(* Logix 5000 project; controller _GigaDiscovery vendor 1 type 14 code 244 rev 35.11; software revision 35.03; part 2 of 23 *)
(* tags used below, declared in another part *)
   Test : DCI_STOP_TEST;

ADD_ON_INSTRUCTION Sfq_Lamp   (* revision 1.0 *)
VAR_INPUT
   Input : BOOL; {required}
END_VAR
VAR_OUTPUT
   LampCoil : BOOL; {access Read Only, visible}
END_VAR
VAR_INPUT
   InputFlt : BOOL; {required}
END_VAR
VAR
   FlsTmr : TIMER := (PRE := 1000); {access None}
END_VAR

ROUTINE Logic   (* ladder *)
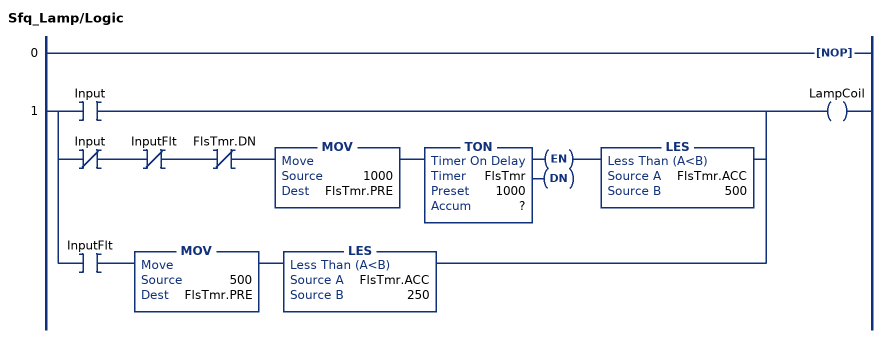
   0: NOP();
   1: [XIC(Input) ,XIO(Input) XIO(InputFlt) XIO(FlsTmr.DN) MOV(1000,FlsTmr.PRE) TON(FlsTmr,?,?) LES(FlsTmr.ACC,500) ,XIC(InputFlt) MOV(500,FlsTmr.PRE) LES(FlsTmr.ACC,250) ]OTE(LampCoil);
END_ROUTINE
END_ADD_ON_INSTRUCTION

ADD_ON_INSTRUCTION Start_AOI   (* revision 1.0 *)
VAR_INPUT
   Start_Ch_1 : BOOL; {required}
   Status_Ch_1 : BOOL; {required}
   Start_Ch_2 : BOOL; {required}
   Status_Ch_2 : BOOL; {required}
   Alarm_Reset : BOOL; {required}
END_VAR
VAR_OUTPUT
   Output : BOOL; {access Read Only, visible}
   Warning : BOOL; {access Read Only, visible}
   Alarm : BOOL; {access Read Only, visible}
   One_Strat_Pb_Pressed : BOOL; {access Read Only}
   Ready : BOOL; {access Read Only}
END_VAR
VAR
   Timer : TIMER[6] := ([0].PRE := 2500, [1].PRE := 2500, [2].PRE := 5000, [3].PRE := 5000, [4].PRE := 5000, [5].PRE := 1000); {access None}
   OS : DINT; {access None}
END_VAR

ROUTINE Logic   (* ladder *)
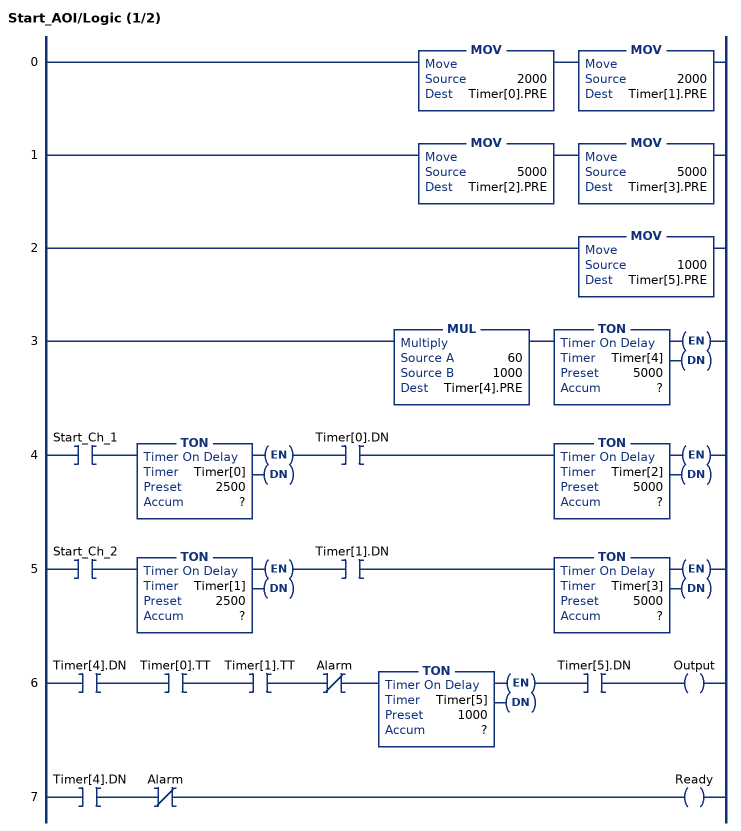
   0: MOV(2000,Timer[0].PRE)MOV(2000,Timer[1].PRE);
   1: MOV(5000,Timer[2].PRE)MOV(5000,Timer[3].PRE);
   2: MOV(1000,Timer[5].PRE);
   3: MUL(60,1000,Timer[4].PRE)TON(Timer[4],?,?);
   4: XIC(Start_Ch_1)TON(Timer[0],?,?)XIC(Timer[0].DN)TON(Timer[2],?,?);
   5: XIC(Start_Ch_2)TON(Timer[1],?,?)XIC(Timer[1].DN)TON(Timer[3],?,?);
   6: XIC(Timer[4].DN)XIC(Timer[0].TT)XIC(Timer[1].TT)XIO(Alarm)TON(Timer[5],?,?)XIC(Timer[5].DN)OTE(Output);
   7: XIC(Timer[4].DN)XIO(Alarm)OTE(Ready);
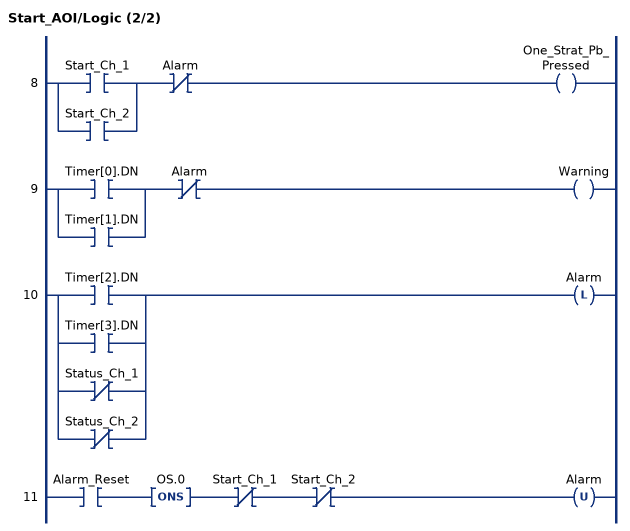
   8: [XIC(Start_Ch_1) ,XIC(Start_Ch_2) ]XIO(Alarm)OTE(One_Strat_Pb_Pressed);
   9: [XIC(Timer[0].DN) ,XIC(Timer[1].DN) ]XIO(Alarm)OTE(Warning);
   10: [XIC(Timer[2].DN) ,XIC(Timer[3].DN) ,XIO(Status_Ch_1) ,XIO(Status_Ch_2) ]OTL(Alarm);
   11: XIC(Alarm_Reset)ONS(OS.0)XIO(Start_Ch_1)XIO(Start_Ch_2)OTU(Alarm);
END_ROUTINE
END_ADD_ON_INSTRUCTION

ADD_ON_INSTRUCTION STD_SCP   (* revision 1.0 *)
VAR_INPUT
   Input : REAL; {required}
   Input_Max : REAL; {required}
   Input_Min : REAL; {required}
END_VAR
VAR_OUTPUT
   Output : REAL; {access Read Only, required}
END_VAR
VAR_INPUT
   Scaled_Max : REAL; {required}
   Scaled_Min : REAL; {required}
END_VAR
VAR
   Rate : REAL;
END_VAR

ROUTINE Logic   (* ladder *)
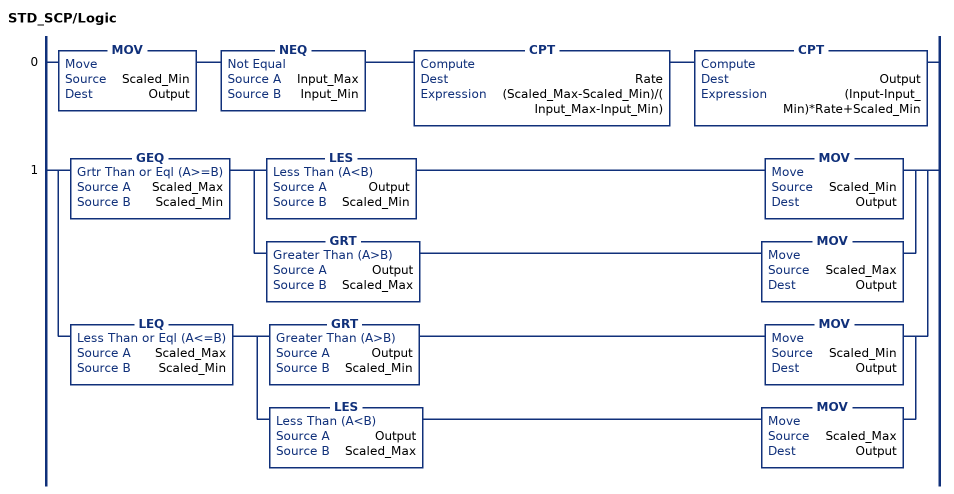
   0: MOV(Scaled_Min,Output)NEQ(Input_Max,Input_Min)CPT(Rate,(Scaled_Max-Scaled_Min)/(Input_Max-Input_Min))CPT(Output,(Input-Input_Min)*Rate+Scaled_Min);
   1: [GEQ(Scaled_Max,Scaled_Min) [LES(Output,Scaled_Min) MOV(Scaled_Min,Output) ,GRT(Output,Scaled_Max) MOV(Scaled_Max,Output) ] ,LEQ(Scaled_Max,Scaled_Min) [GRT(Output,Scaled_Min) MOV(Scaled_Min,Output) ,LES(Output,Scaled_Max) MOV(Scaled_Max,Output) ] ];
END_ROUTINE
END_ADD_ON_INSTRUCTION

ADD_ON_INSTRUCTION Valve_2_pos_monostable   (* revision 1.0 *)
VAR_INPUT
   I_Enable : BOOL; {required}
   FeedBack_Type : BOOL; {required}   // 0 = Equivalent 1 = Reverse
   Discrepancy_Time : DINT; {access None, required}
   I_FeedBack_Data : BOOL; {required}
   I_FeedBack_Status : BOOL; {required}
   I_Output_Status : BOOL; {required}
   I_Fault_Reset : BOOL; {required}
END_VAR
VAR_OUTPUT
   FP : BOOL; {access Read Only, visible}
   O1 : BOOL; {access Read Only, visible}
   O_ERR : DINT; {access Read Only}
END_VAR
VAR
   ON_Delay_Control : TIMER; {access None}
   OFF_Delay_Control : TIMER; {access None}
   Fault_Condiction : BOOL; {access None}
   ONS : BOOL; {access None}
END_VAR

ROUTINE Logic   (* ladder *)
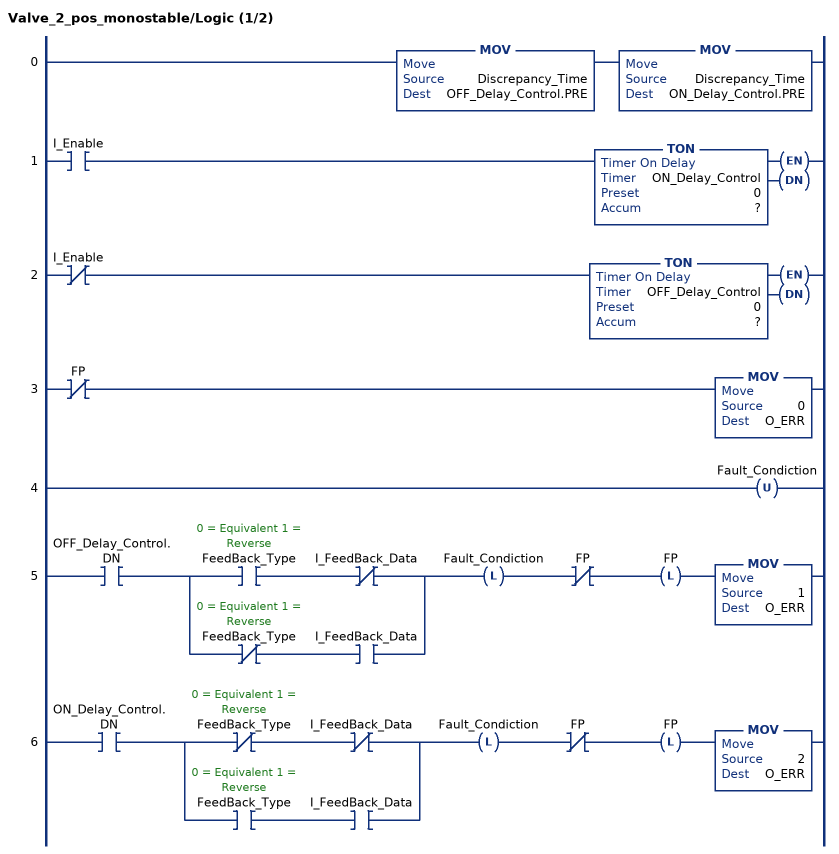
   0: MOV(Discrepancy_Time,OFF_Delay_Control.PRE)MOV(Discrepancy_Time,ON_Delay_Control.PRE);
   1: XIC(I_Enable)TON(ON_Delay_Control,?,?);
   2: XIO(I_Enable)TON(OFF_Delay_Control,?,?);
   3: XIO(FP)MOV(0,O_ERR);
   4: OTU(Fault_Condiction);
   5: XIC(OFF_Delay_Control.DN)[XIC(FeedBack_Type) XIO(I_FeedBack_Data) ,XIO(FeedBack_Type) XIC(I_FeedBack_Data) ]OTL(Fault_Condiction)XIO(FP)OTL(FP)MOV(1,O_ERR);
   6: XIC(ON_Delay_Control.DN)[XIO(FeedBack_Type) XIO(I_FeedBack_Data) ,XIC(FeedBack_Type) XIC(I_FeedBack_Data) ]OTL(Fault_Condiction)XIO(FP)OTL(FP)MOV(2,O_ERR);
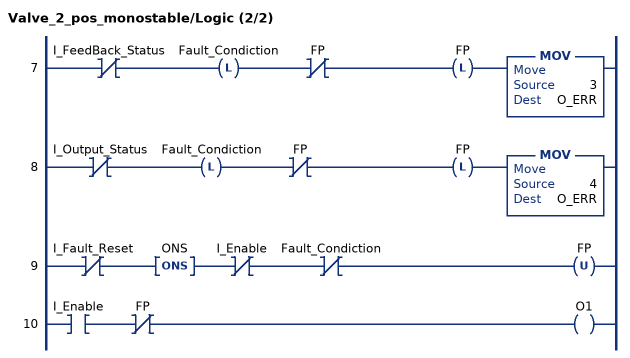
   7: XIO(I_FeedBack_Status)OTL(Fault_Condiction)XIO(FP)OTL(FP)MOV(3,O_ERR);
   8: XIO(I_Output_Status)OTL(Fault_Condiction)XIO(FP)OTL(FP)MOV(4,O_ERR);
   9: XIO(I_Fault_Reset)ONS(ONS)XIO(I_Enable)XIO(Fault_Condiction)OTU(FP);
   10: XIC(I_Enable)XIO(FP)OTE(O1);
END_ROUTINE
END_ADD_ON_INSTRUCTION

VAR_GLOBAL   (* controller tags *)
   Acc_Time : REAL := 0.5;   // T2 Region 2
   All_Rack_Closed_Mem : BOOL := 1;
   All_Rack_Left_Sensor_FP_OFF : BOOL := 1;
   All_Rack_Left_Sensor_O1_OFF : BOOL;
   All_Rack_Right_Sensor_FP_OFF : BOOL := 1;
   All_Rack_Right_Sensor_O1_OFF : BOOL;
   All_Rack_Sensor_OFF : BOOL;
   All_RESTRAINTS_Opened : BOOL;
   Analog_Input_Pos_6 : REAL[8] := ([0] := 0.0061035156, [2] := -0.025939941, [4] := -0.025939941, [6] := -0.0289917);
        [0]   // Lettura tensione Motori 1 - 3 Pilone
        [1]   // Lettura Corrente Motori 1 - 3 Pilone
        [2]   // Lettura tensione Motori 2 - 4 Pilone
        [3]   // Lettura Corrente Motori 2 - 4 Pilone
        [6]   // Lettura tensione Motori 5 - 6 Pilone
        [7]   // Lettura Corrente Motori 5 - 6 Pilone
        [4]   // Lettura tensione Motore Gondola
        [5]   // Lettura Corrente Motore Gondola
   Analog_Output_Pos_5 : REAL[8] := ([4] := 10000.0);
        [4]   // Gondola Torque Limit
        [5]   // Gondola Speed Reference
   Angle_at_Full_Load : REAL := 12.0;
   Angle_at_min_Load : REAL := 14.0;
   Angle_Controll_S_Curve : S_Curve_Calc := (Jerk_Time := 0.5, Accel_Time := 1.0, Jerk_Rate := 300.0, Accel_Rate := 150.0);
   AngleContrl : REAL := 77.39982;
   Auto_Cycle_Step : DINT := 1;
   auto_manual : TIMER := (PRE := 2000);
   Automatic_Cycle_DB : Auto_Cycle[6] := ([1].Pylon_Angle := 120, [1].Cycle_Time_min := 2, [1].Cycle_Time_sec := 25, [1].Gondola_Speed[0] := 20, [1].Gondola_Speed[1] := 70, [1].Gondola_Speed[2] := -75, [1].Gondola_Speed[3] := 50, [1].Gondola_Time[1] := 60, [1].Gondola_Time[2] := 50, [1].Gondola_Time[3] := 20, [2].Pylon_Angle := 90, [2].Cycle_Time_min := 1, [2].Cycle_Time_sec := 50, [2].Gondola_Speed[1] := 50, [2].Gondola_Speed[2] := -75, [2].Gondola_Speed[3] := 50, [2].Gondola_Time[0] := 90, [2].Gondola_Time[1] := 60, [2].Gondola_Time[2] := 50, [2].Gondola_Time[3] := 20, [3].Pylon_Angle := 75, [3].Cycle_Time_min := 1, [3].Cycle_Time_sec := 30, [3].Gondola_Speed[1] := 50, [3].Gondola_Speed[2] := -50, [3].Gondola_Speed[3] := -100, [3].Gondola_Time[1] := 60, [3].Gondola_Time[2] := 60, [4].Pylon_Angle := 45, [4].Cycle_Time_min := 1, [4].Cycle_Time_sec := 20, [4].Gondola_Speed[1] := 50, [4].Gondola_Speed[2] := -50, [4].Gondola_Time[1] := 60, [4].Gondola_Time[2] := 50, [5].Pylon_Angle := 20, [5].Cycle_Time_min := 10, [5].Gondola_Time[1] := 60);
   Automatic_E_Stop_Cl_0 : DINT := -1;
   Automatic_E_Stop_Cl_1 : DINT := -1;
   Braking_Torque_Lim : REAL := 20.0;
   CCW_OS_Direction_1 : BOOL;
   CCW_OS_Direction_2 : BOOL;
   Clock : DINT := -1934744665;   // Base tempi 10 milli sec
        .8   // 5,12 sec
        .6   // 1280 milli sec
        .0   // 20 milli sec
        .7   // 2560 milli sec
        .3   // 160 milli sec
        .1   // 40 milli sec
        .2   // 80 milli sec
        .4   // 320 milli sec
        .5   // 640 milli sec
   Clock_1_Hz : BOOL;   // SL Clock 1 Hz 0.5 sec OFF 0.5 sec ON
   Clock_4_Hz : BOOL := 1;   // SL Clock 4 Hz 0.125 sec OFF 0.125 sec ON
   Close_Platform_Autocycle_Pylon : BOOL;
   Compressor_Pressure_OK : BOOL := 1;
   CROUT_Air_Compressor : UDT_CROUT := (CROUT.Actuate := 1, CROUT.InputStatus := 1, CROUT.OutputStatus := 1, CROUT.FeedbackReactionTime := 500, CROUT.O1 := 1, CROUT.O2 := 1);   // Compressor Command -Q18101E
   Current_TimeInStation : DINT;
   CurrentLimit : DINT := 100;
   CW_OS_Direction_1 : BOOL;
   CW_OS_Direction_2 : BOOL;
   Cycle_End_Timer : TIMER := (PRE := 60000);
   Cycle_Time : TIMER := (PRE := 145000);
   Cycle_Timing : TIMER := (PRE := 600000);
   CycleOver : BOOL;
   DC_Field_Motor_7 : UDT_CROUT := (CROUT.Feedback1 := 1, CROUT.Feedback2 := 1, CROUT.InputStatus := 1, CROUT.OutputStatus := 1, CROUT.FeedbackReactionTime := 500, Timer.PRE := 100, Timer.ACC := 100);   // DC Field Motor 7 Gondola Contactor -Q16101E -Q16103E
   DC_Field_Pylon_Motors : UDT_CROUT := (CROUT.Feedback1 := 1, CROUT.Feedback2 := 1, CROUT.InputStatus := 1, CROUT.OutputStatus := 1, CROUT.FeedbackReactionTime := 500, Timer.PRE := 100, Timer.ACC := 120);   // DC Field Pylon Motors Contactor -Q10101E -Q10103E
   Direction : BOOL := 1;   // 1 = Spinta CW 0 = Spinta CCW
   E_Stop2_Test_Request : BOOL;
   E_Stop_Secondary_Test_Ok : BOOL := 1;
   E_Stop_Test_Request : BOOL;
   Echo_HMI_Modify_Auto_Cycle_Ptr : DINT := 1;
   Emergencies_CL0 : DINT[8];
        [5].0   // CYCLE - Field Contactor Feedback Motor 1-2 Fault -Q10101E -Q10103E -Q10202G
        [5].17   // CYCLE - Motor 1-2 Field contactor -Q10101E -Q10103E -Q10202G remain ON
        [2].4   // PLATFORM - Platform not opened -B22501J ... -B22807J -B22501B
        [5].26   // Valve Proof Test Failed - Open/Close Platform Valves do not work correctly
        [1].8   // PLATFORM - Pressure in Pilot Valve Line with Valve OFF -S22006B
        [5].19   // CYCLE - Motor 7 Field contactor -Q16101E -Q16103E -Q16202G remain ON
        [1].0   // PLATFORM - Pressure Switch -21504B Unespected remains ON
        [0].10   // +RCC_GSG Temperature -S62110G
        [5].28   // Valve Proof Test Failed - Platform moved during test
        [5].29   // Valve Proof Test Failed - Platform moved during test
        [5].5   // CYCLE - Field Contactor Feedback Motor 7 Fault -Q16101E -Q16103E -Q16202G
        [0].11   // +RCC_GSG Temperature -S64110G
        [0].3   // +RCC_GSA Temperature OK -S50410G
        [1].1   // PLATFORM - Pressure Switch -21504B Unespected remains OFF
        [4].1   // PYLON - Overlimit sensor fault -A26510I
        [0].4   // +GMB_RCC1 Temperature OK -S40103E
        [2].3   // PLATFORM - Platform not closed -B23501J ... -B23807J -B23501F
        [2].7   // PLATFORM - Platform not closed -B23501J ... -B23807J -B23501F
        [1].5   // PLATFORM - Pressure Switch -21504B Unespected remains ON
        [5].10   // CYCLE - Motor 5-6 Converter remain ON
        [5].27   // Valve Proof Test Failed - Pressure in Line with Main Valve OFF
        [2].0   // PLATFORM - Pressure Switch -21511B Unespected remains ON
        [4].2   // Gondola Overspeed from Sensor -B40002I
        [4].4   // Gondola Overspeed from Sensor -B40007I
        [5].6   // CYCLE - Motor 5-6 Converter not Active
        [2].1   // PLATFORM - Pressure Switch -21511B Unespected remains ON
        [5].11   // CYCLE - Motor 1-2 Converter remain ON
        [1].6   // PLATFORM -Platform not open -B22501J ... -B22807J -B22501B
        [5].12   // CYCLE - Motor 3-4 Converter remain ON
        [5].14   // CYCLE - Motor 1-2 Converter remain ON
        [2].2   // PLATFORM - Pressure Switch -21510B Unespected remains ON
        [2].5   // PLATFORM - Pressure Switch -21507B Unespected remains ON
        [2].6   // PLATFORM - Pressure Switch -21511B Unespected remains ON
        [5].15   // CYCLE - Motor 3-4 Converter remain ON
        [5].21   // CYCLE - Motor 5-6 Converter remain ON
        [0].0   // Restraints Right Pressure Switch remains on
        [5].20   // OCC2 Control Disable Input Fault Page 310
        [5].25   // Valve Proof Test Failed - No pressure with Main Valve ON
        [5].24   // CYCLE - Motor 5-6 Converter not Ready
        [5].9   // CYCLE - Motor 7 Converter not Active
        [1].10   // Platform main valve B21902I Fault
        [5].7   // CYCLE - Motor 1-2 Converter not Active
        [4].3   // PYLON - Overlimit sensor hit -A26510I
        [1].7   // PLATFORM - Pilot Valve Line has not pressure -S22006B
        [0].7   // +RCC_GSD Temperature -S56110G
        [5].1   // CYCLE - Motor 1-2 Converter not Ready
        [5].8   // CYCLE - Motor 3-4 Converter not Active
        [5].13   // CYCLE - Motor 7 Converter remain ON
        [5].16   // CYCLE - Motor 7 Converter remain ON
        [5].2   // CYCLE - Motor 3-4 Converter not Ready
        [1].2   // PLATFORM - Platform not closed
        [0].1   // Restraints Left Pressure Switch remains on
        [1].3   // PLATFORM - Platform not opened
        [0].8   // +RCC_GSE Temperature -S58110G
        [4].0   // Pylon Overspeed B26202A B26206A
        [0].12   // Retraints Opened During ProofTest
        [5]   // Automatic cycle
        [1].4   // PLATFORM - Not used
        [0].9   // +RCC_GSF Temperature -S60110G
        [5].3   // CYCLE - Motor 7 Converter not Ready
        [0].5   // +RCC_GSB Temperature OK -S52110G
        [0].6   // +RCC_GSC Temperature OK -S54110G
        [0].2   // Restraints Not Closed
        [5].4   // CYCLE - Start Contactors Failed to Actuate -Q
        [1].9   // Compressor Command -Q18101E Contactor Fault
   Emergencies_CL1 : DINT[14];
        [5].21   // LAPBARS - SECTOR C Seat 11-15 Opened During Cycle -B55001J -B55007J -B55101J -B55107J -B55201J
        [5].19   // LAPBARS - SECTOR A Seat 1-5 Opened During Cycle -B51001J -B51007J -B51101J -B51107J -B51201J
        [10].0   // Platform Line Minimum Pressure Switch -S21511B Signal missing during Start Cycle
        [5].20   // LAPBARS - SECTOR B Seat 6-10 Opened During Cycle -B53001J -B53007J -B53101J -B53107J -B53201J
        [5].22   // LAPBARS - SECTOR D Seat 16-20 Opened During Cycle -B57001J -B57007J -B57101J -B57107J -B57201J
        [3].10   // MCC - Gondola Drive Enable Contactors Feeback Fault -Q16105E -Q16107E
        [5].8   // GATE OPERATOR 4 RFID SENSOR - EAC-5 -B24803J Opened during cycle
        [3].1   // MCC - Pylon Start Drive 1-2 Contactors Feedback Fault -Q9002E -Q9004E
        [5].2   // PLATFORM - Close Sensor Discrepancy Fault -B22501J ... -B22807J -B22501B
        [10].1   // Platform Proof Test Unlock Line Pressure Switch -S22006B Signsl missing
        [2].3   // OCC - Start Enable and Start Button Fault -S30401F -S30403F
        [3].4   // MCC - DC Motor 7 Gondola Contactor Feedabck fault -Q16101E -Q16103E
        [5].23   // LAPBARS - SECTOR E Seat 21-25 Opened During Cycle -B59001J -B59007J -B59101J -B59107J -B59201J
        [10].2   // Platform Proof Test Open Main Valve Limit Switch -B21905I Signsl missing
        [10].3   // Platform Proof Test Opened RFID Series -Q23801J -Q23807J Signsl missing
        [7].2   // LAPBARS - SECTOR B Unlock Right Feedback Fault, Y10202F
        [3].9   // Pylon Start Drive 5 - 6 Contactors -Feedback Fault Q9009E -Q9011E4 -Q14202G -Q14202G
        [3].3   // MCC - Pylon Start Drive 3-4 Contactors Feedback Fault -Q9005E -Q9007E
        [3].27   // -S28507F RESTRAINTS RELEASE UNLOCK -RUN- LOCK RESTRAINTS selector Fault
        [7].10   // LAPBARS - SECTOR F Unlock Right Feedback Fault, Y12202F
        [7].12   // LAPBARS - SECTOR G Unlock Right Feedback Fault, Y12702F
        [7].11   // LAPBARS - SECTOR F Unlock Left Feedback Fault, Y12205F
        [5].24   // LAPBARS - SECTOR F Seat 26-30 Opened During Cycle -B61001J -B61007J -B61101J -B61107J -B61201J
        [3].2   // MCC - DC Motor 1-2 Contactor Feedabck fault -Q10101E -Q10103E
        [5].25   // LAPBARS - SECTOR G Seat 31-35 Opened During Cycle -B63001J -B63007J -B63101J -B63107J -B63201J
        [5].26   // LAPBARS - SECTOR H Seat 36-40 Opened During Cycle -B65001J -B65007J -B65101J -B65107J -B65201J
        [7].13   // LAPBARS - SECTOR G Unlock Left Feedback Fault, Y12705F
        [7].4   // LAPBARS - SECTOR C Unlock Right Feedback Fault, Y10702F
        [7].0   // LAPBARS - SECTOR A Unlock Right Feedback Fault, Y9702F
        [4].16   // LAPBARS - SECTOR A key enable signal fault -S27802F
        [7].3   // LAPBARS - SECTOR B Unlock Left Feedback Fault, Y10205F
        [7].6   // LAPBARS - SECTOR D Unlock Right Feedback Fault, Y11202F
        [4].17   // LAPBARS - SECTOR B key enable signal fault -S27806F
        [7].5   // LAPBARS - SECTOR C Unlock Left Feedback Fault, Y10705F
        [7].7   // LAPBARS - SECTOR D Unlock Left Feedback Fault, Y11205F
        [4].18   // LAPBARS - SECTOR C key enable signal fault -S27902F
        [7].8   // LAPBARS - SECTOR E Unlock Right Feedback Fault, Y11702F
        [7].9   // LAPBARS - SECTOR E Unlock Left Feedback Fault, Y11705F
        [4].19   // LAPBARS - SECTOR D key enable signal fault -S27906F
        [3].0   // OCC2 Allow Main CONFIRM -S28602F Stucked Close
        [0].17   // GONDOLA GMB - Mudule Fault K39001C
        [5].3   // PLATFORM - Open Sensor Discrepancy Fault -B23501J...-B23807J -B23501F
        [0].18   // GONDOLA GMB - Mudule Fault K39002C
        [7].14   // LAPBARS - SECTOR H Unlock Right Feedback Fault, Y13202F
        [0].19   // GONDOLA GMB - Mudule Fault K39003C
        [4].0   // LAPBARS - SECTOR A Open during cycle
        [7].15   // LAPBARS - SECTOR H Unlock Right Feedback Fault, Y13205F
        [8].11   // LAPBARS - SECTOR A Seat 1 Opened During Cycle -B51001J
        [0].24   // GONDOLA GSA - Mudule Fault K39501C
        [8].20   // LAPBARS - SECTOR B Seat 10 Opened During Cycle -B53201J
        [0].25   // GONDOLA GSA - Mudule Fault K39502C
        [4].1   // LAPBARS - SECTOR B Open during cycle
        [0].26   // GONDOLA GSA - Mudule Fault K39503C
        [0].27   // GONDOLA GSA - Mudule Fault K39504C
        [6].0   // Pylon - Fan Contactors Feedback Fault - Not all closed Pag.94
        [8].12   // LAPBARS - SECTOR A Seat 2 Opened During Cycle -B51007J
        [2].7   // Entry Gate selector turned during cycle
        [2].8   // Exit Gate selector turned during cycle
        [6].1   // Pylon - Fan Contactors Feedback Fault - Not all open Pag.94
        [5].9   // GATE ENTER (G01) -B25204I Opened during cycle
        [8].13   // LAPBARS - SECTOR A Seat 3 Opened During Cycle -B51101J
        [9].10   // LAPBARS - SECTOR G Seat 32 Opened During Cycle -B63007J
        [0].28   // GONDOLA GSB - Mudule Fault K52001C
        [4].20   // LAPBARS - SECTOR E key enable signal fault -S28002F
        [8].14   // LAPBARS - SECTOR A Seat 4 Opened During Cycle -B51107J
        [8].21   // LAPBARS - SECTOR C Seat 11 Opened During Cycle -B55001J
        [8].22   // LAPBARS - SECTOR C Seat 12 Opened During Cycle -B55007J
        [8].23   // LAPBARS - SECTOR C Seat 13 Opened During Cycle -B55101J
        [3].11   // MCC - Gondola Motor Power Supply Fuses Blown -F16002F -F16003F
        [9].11   // LAPBARS - SECTOR G Seat 33 Opened During Cycle -B63101J
        [0].29   // GONDOLA GSB - Mudule Fault K52002C
        [8].15   // LAPBARS - SECTOR A Seat 5 Opened During Cycle -B51201J
        [8].16   // LAPBARS - SECTOR B Seat 6 Opened During Cycle -B53001J
        [9].12   // LAPBARS - SECTOR G Seat 34 Opened During Cycle -B63107J
        [9].0   // LAPBARS - SECTOR E Seat 22 Opened During Cycle -B59007J
        [8].24   // LAPBARS - SECTOR C Seat 14 Opened During Cycle -B55107J
        [0].30   // GONDOLA GSB - Mudule Fault K52003C
        [8].25   // LAPBARS - SECTOR C Seat 15 Opened During Cycle -B55201J
        [4].21   // LAPBARS - SECTOR F key enable signal fault -S28006F
        [8].26   // LAPBARS - SECTOR D Seat 16 Opened During Cycle -B57001J
        [5].5   // PLATFORM - Platform Open and Close at same time
        [1].10   // MCC - Input Fault K20801C
        [4].2   // LAPBARS - SECTOR C Open during cycle
        [1].12   // OCC - Input Fault K30001C
        [8].27   // LAPBARS - SECTOR D Seat 17 Opened During Cycle -B57007J
        [1].13   // OCC - Input Fault K30002C
        [8].28   // LAPBARS - SECTOR D Seat 18 Opened During Cycle -B57101J
        [0].31   // GONDOLA GSB - Mudule Fault K52004C
        [2].0   // OCC - Lapbars selector fault -S30505F
        [1].14   // OCC - Input Fault K30003C
        [2].10   // GONDOLA GSB - Mudule Fault K54001C
        [2].11   // GONDOLA GSB - Mudule Fault K54002C
        [2].12   // GONDOLA GSB - Mudule Fault K52003C
        [2].13   // GONDOLA GSB - Mudule Fault K52004C
        [7].16   // LAPBARS - SECTOR A Close Sensor Discrepancy Fault
        [7].17   // LAPBARS - SECTOR B Close Sensor Discrepancy Fault
        [1].15   // MCC - Input Fault K20803C
        [1].16   // GSA - Output Fault K50004C
        [8].29   // LAPBARS - SECTOR D Seat 19 Opened During Cycle -B57107J
        [8].30   // LAPBARS - SECTOR D Seat 20 Opened During Cycle -B57201J
        [2].14   // GONDOLA GSD - Mudule Fault K56001C
        [2].15   // GONDOLA GSD - Mudule Fault K56002C
        [7].19   // LAPBARS - SECTOR D Close Sensor Discrepancy Fault
        [2].16   // GONDOLA GSD - Mudule Fault K56003C
        [8].31   // LAPBARS - SECTOR E Seat 21 Opened During Cycle -B59001J
        [2].5   // OCC- LockOut Motion Component Fault -Q31203E
        [6].7   // Home Sensor Speed Check -B40002I Fault
        [5].0   // PLATFORM - Main Valve Feedback Fault -B21902I
        [3].29   // OCC2 - E-Stop Pressed -S28502F
        [3].28   // OCC - E-Stop Pressed -S30301F
        [4].3   // LAPBARS - SECTOR D Open during cycle
        [7].20   // LAPBARS - SECTOR E Close Sensor Discrepancy Fault
        [9].1   // LAPBARS - SECTOR E Seat 23 Opened During Cycle -B59101J
        [8].17   // LAPBARS - SECTOR B Seat 7 Opened During Cycle -B53007J
        [7].18   // LAPBARS - SECTOR C Close Sensor Discrepancy Fault
        [8].3   // GATE 4 OPERATOR RFID SENSOR - MOP -B25404J Fault
        [0].0   // MCC - Mudule Fault K20501C
        [0].1   // MCC - Mudule Fault K20502C
        [6].8   // Home Sensor Speed Check -B40007I Fault
        [4].4   // LAPBARS - SECTOR E Open during cycle
        [4].5   // LAPBARS - SECTOR F Open during cycle
        [2].17   // GONDOLA GSD - Mudule Fault K56004C
        [2].18   // GONDOLA GSE - Mudule Fault K58001C
        [2].19   // GONDOLA GSE - Mudule Fault K58002C
        [9].2   // LAPBARS - SECTOR E Seat 24 Opened During Cycle -B59107J
        [9].3   // LAPBARS - SECTOR E Seat 25 Opened During Cycle -B59201J
        [9].8   // LAPBARS - SECTOR F Seat 30 Opened During Cycle -B61201J
        [9].13   // LAPBARS - SECTOR G Seat 35 Opened During Cycle -B63201J
        [1].23   // GSB - Output Fault K52004C
        [7].21   // LAPBARS - SECTOR F Close Sensor Discrepancy Fault
        [0].2   // MCC - Mudule Fault K20503C
        [2].20   // GONDOLA GSE - Mudule Fault K58003C
        [1].26   // GSC - Output Fault K52004C
        [7].22   // LAPBARS - SECTOR G Close Sensor Discrepancy Fault
        [9].14   // LAPBARS - SECTOR H Seat 36 Opened During Cycle -B65001J
        [2].21   // GONDOLA GSE - Mudule Fault K58004C
        [2].31   // GSD - Output Fault K56004C
        [2].22   // GONDOLA GSF - Mudule Fault K60001C
        [4].22   // LAPBARS - SECTOR G key enable signal fault -S28102F
        [8].18   // LAPBARS - SECTOR B Seat 8 Opened During Cycle -B53101J
        [8].19   // LAPBARS - SECTOR B Seat 9 Opened During Cycle -B53107J
        [6].2   // PYLON - Home position Ch1 Fault -B26002I
        [6].3   // PYLON - Home position Ch2 Fault -B26007I
        [9].15   // LAPBARS - SECTOR H Seat 37 Opened During Cycle -B65007J
        [0].20   // GONDOLA GMB Fault K39004C
        [9].4   // LAPBARS - SECTOR F Seat 26 Opened During Cycle -B61001J
        [2].23   // GONDOLA GSF - Mudule Fault K60002C
        [0].22   // GSC - Input Fault K54003C
        [0].23   // GSA - Input Fault K50003C
        [5].10   // GATE EXIT (G05) -B25304I Opened during cycle
        [2].24   // GONDOLA GSF - Mudule Fault K60003C
        [0].3   // MCC - Mudule Fault K20504C
        [9].16   // LAPBARS - SECTOR H Seat 38 Opened During Cycle -B65101J
        [9].17   // LAPBARS - SECTOR H Seat 39 Opened During Cycle -B65107J
        [2].25   // GONDOLA GSF - Mudule Fault K60004C
        [0].4   // MCC - Mudule Fault K20505C
        [2].26   // GONDOLA GSG - Mudule Fault K62001C
        [3].13   // GSE - Output Fault K58004C
        [2].27   // GONDOLA GSG - Mudule Fault K62002C
        [9].18   // LAPBARS - SECTOR H Seat 40 Opened During Cycle -B65201J
        [4].6   // LAPBARS - SECTOR G Open during cycle
        [2].28   // GONDOLA GSG - Mudule Fault K62003C
        [0].5   // MCC - Mudule Fault K20506C
        [4].7   // LAPBARS - SECTOR H Open during cycle
        [0].6   // MCC - Mudule Fault K20507C
        [0].7   // MCC - Mudule Fault K20508C
        [0].8   // MCC - Mudule Fault K20509C
        [0].9   // MCC - Module Fault K20518C
        [3].17   // GSF - Output Fault K60004C
        [3].21   // GSG - Output Fault K62004C
        [9].5   // LAPBARS - SECTOR F Seat 27 Opened During Cycle -B61007J
        [2].29   // GONDOLA GSG - Mudule Fault K62004C
        [3].25   // GSH - Output Fault K64004C
        [4].8   // LAPBARS - Sector Enabled A-B
        [4].23   // LAPBARS - SECTOR H key enable signal fault -S28106F
        [1].20   // GSB - Input Fault K52001C
        [1].21   // GSB - Input Fault K52002C
        [1].22   // GSB - Input Fault K52003C
        [4].10   // LAPBARS - Sector Enabled C-D
        [1].24   // GSA - Input Fault K50001C
        [6].4   // Zero Set Sensor Missing B11201A
        [4].9   // LAPBARS - Sector Enabled B-C
        [9].6   // LAPBARS - SECTOR F Seat 28 Opened During Cycle -B61101J
        [2].30   // GONDOLA GSH - Mudule Fault K62001C
        [4].11   // LAPBARS - Sector Enabled D-E
        [1].25   // GSA - Input Fault K50002C
        [7].1   // LAPBARS - SECTOR A Unlock Left Feedback Fault, Y9705F
        [1].27   // GSC - Input Fault K54001C
        [9].7   // LAPBARS - SECTOR F Seat 29 Opened During Cycle -B61107J
        [9].9   // LAPBARS - SECTOR G Seat 31 Opened During Cycle -B63001J
        [1].28   // GSC - Input Fault K54002C
        [2].1   // Alarm OCC temperature OK -S31003E
        [7].23   // LAPBARS - SECTOR H Close Sensor Discrepancy Fault
        [2].6   // OCC- FootPedal Component Fault -S30901F
        [1].29   // GSD - Input Fault K56001C
        [5].1   // Time Out Open Platform cycle
        [1].30   // GSD - Input Fault K56002C
        [4].12   // LAPBARS - Sector Enabled E-F
        [3].5   // OCC Aut/Man Selector Fault S30801F
        [0].11   // MCC - Mudule Fault K20801B
        [1].31   // GSD - Input Fault K56003C
        [0].12   // MCC - Mudule Fault K30001B
        [4].13   // LAPBARS - Sector Enabled F-G
        [2].9   // Operator Gate selector turned during cycle
        [0].13   // MCC - Mudule Fault K30002B
        [4].14   // LAPBARS - Sector Enabled G-H
        [4].15   // LAPBARS - Sector Enabled H-A
        [0].14   // OCC - Mudule Fault K30003B
        [4].25   // LAPBARS - Main Air Line Pressure Missing
        [0].15   // MCC - Mudule Fault K20802B
        [0].16   // MCC - Mudule Fault K20803B
        [1].11   // MCC - Output Fault K20802C
        [1].17   // RCC 1 - Input Fault K39001C
        [3].26   // UPS MCC -T6603B Alarm
        [2].2   // OCC - E-Stop Fault -S30301F
        [1].18   // RCC 1 - Input Fault K39002C
        [1].19   // RCC 1 - Input Fault K39003C
        [0]   // Communication
        [2].4   // OCC 2 - E-Stop Fault -S28502F
        [3].14   // GSF - Input Fault K60001C
        [3].15   // GSF - Input Fault K60002C
        [3].16   // GSF - Input Fault K60003C
        [8].2   // GATE ENTER (G01) -B25204I Fault
        [3].6   // GSE - Input Fault K58001C
        [3].18   // GSG - Input Fault K62001C
        [3].12   // UPS RCC -T37603B Alarm
        [3].7   // GSE - Input Fault K58002C
        [1].0   // MCC - Input Fault K20501C
        [1].1   // MCC - Input Fault K20502C
        [1].2   // MCC - Input Fault K20503C
        [1].3   // MCC - Input Fault K20504C
        [1].4   // MCC - Input Fault K20505C
        [1].5   // MCC - Input Fault K20506C
        [1].6   // MCC - Input Fault K20507C
        [1].7   // MCC - Input Fault K20508C
        [1].8   // MCC - Input Fault K20509C
        [1]   // I/O Status
        [1].9   // MCC - Input Fault K20518C
        [3].19   // GSG - Input Fault K62002C
        [3].20   // GSG - Input Fault K62003C
        [3].22   // GSH - Input Fault K64001C
        [3].23   // GSH - Input Fault K64002C
        [3].8   // GSE - Input Fault K58003C
        [3].24   // GSH - Input Fault K64003C
        [6].6   // Home Sensor Speed Stack
        [8].1   // GATE EXIT (G05) -B25304I
        [5].6   // PLATFORM - Platform not openend during cycle
        [6].5   // PYLON - Brake command Feedbak Fault -Q10801E
        [8].0   // GATE 4 RFID SENSOR - EAC-5 -B24803J Fault
        [4].24   // LAPBARS - Main valve command Fault -B45001I
   Emergencies_Std_CL0 : DINT[8];
        [0].15   // Code 0.15 Termic Probe Gondola Motor 5 B6007C Rif. KA6007H
        [0].9   // Pylon Angle Overlimit Alarm by Encoder
        [2].14   // Code 2.14 Dig Out 1 DC Converter Mot 1_3 T608C Rif. FIELD LOSS